// TIA Portal project "pb_slave_test_ZASI_V18" (V18)

(* hardware
DEVICE "S7-1200 station_1"  S7-1200 Station
   slot 0: "Rack_0"  S7-1200 Rack  Rack  V1.0
   slot 1: "PLC_1"  CPU 1212C AC/DC/Rly  6ES7 212-1BE40-0XB0  V4.3
   slot 101: "CM 1243-5"  CM 1243-5  6GK7 243-5DX30-0XE0  V1.3
DEVICE "HMI_1"  KTP700 Basic PN
   slot 0: "HMI_1"  KTP700 Basic PN  6AV2 123-2GB03-0AX0  15.1.0.0
   slot 1: "HMI_RT_1"  KTP700 Basic PN  6AV2 123-2GB03-0AX0  15.1.0.0
   slot 5: "HMI_1.IE_CP_1"  PROFINET Interface  15.0.1.0
      slot 1: "PROFINET Interface_1"  PROFINET Interface
         slot 1: "Port_1"  Port
DEVICE "GSD device_1"  GSD.Device
   slot 0: "Rack_0"  Rail
*)

// ===== PLC "PLC_1"  CPU 1212C AC/DC/Rly =====

VAR_GLOBAL   // PLC tag table "Default tag table"
   "Tag_2" AT %I0.0 : Bool;
   "Tag_1" AT %Q0.0 : Bool;
   "ProfiOut" AT %Q1.0 : "DataRange";
   "System_Byte" AT %MB1 : Byte;
   "FirstScan" AT %M1.0 : Bool;
   "DiagStatusUpdate" AT %M1.1 : Bool;
   "AlwaysTRUE" AT %M1.2 : Bool;
   "AlwaysFALSE" AT %M1.3 : Bool;
   "Clock_Byte" AT %MB0 : Byte;
   "Clock_10Hz" AT %M0.0 : Bool;
   "Clock_5Hz" AT %M0.1 : Bool;
   "Clock_2.5Hz" AT %M0.2 : Bool;
   "Clock_2Hz" AT %M0.3 : Bool;
   "Clock_1.25Hz" AT %M0.4 : Bool;
   "Clock_1Hz" AT %M0.5 : Bool;
   "Clock_0.625Hz" AT %M0.6 : Bool;
   "Clock_0.5Hz" AT %M0.7 : Bool;
   "Length" AT %MD100 : DInt;
   "Length_of_buht" AT %MD104 : DInt;
   "Length_of_buht_current" AT %MD108 : DInt;
   "Velocity" AT %MD112 : DInt;
   "ProfiIn" AT %I1.0 : "DataRange";
   "Dm_pb" AT %ID35 : DWord;
   "Dx_pb" AT %ID39 : UDInt;
   "Dy_pb" AT %ID43 : UDInt;
   "Cx_pb" AT %ID47 : UDInt;
   "Cy_pb" AT %ID51 : UDInt;
   "Error_pb" AT %IB55 : Byte;
   "L_all" AT %ID1 : DInt;
   "set_buht" AT %ID9 : UDInt;
   "L_buht" AT %ID5 : DInt;
   "vel" AT %ID13 : UDInt;
   "Tag_3" AT %QB0 : Byte;
   "Tag_4" AT %QD3 : DInt;
   "ZASI_pb_write_data_addr" AT %QB1 : Byte;
   "Tag_6" AT %QD4 : DInt;
   "Tag_7" AT %QD2 : DInt;
   "ustavka_out" AT %QW6 : Word;
   "proboy" AT %QW4 : Word;
   "reset_length" AT %QB3 : Byte;
   "Ustavka" AT %IW9 : UInt;
   "Voltage" AT %IW13 : UInt;
   "Hi_on" AT %QW2 : UInt;
END_VAR

VAR_GLOBAL   // PLC tag table "global_tags"
   "need_write" AT %M110.0 : Bool;
   "write_addr" AT %MB111 : Byte;
   "new_val" AT %MB112 : Byte;
   "dev_addr" AT %MB113 : Byte;
END_VAR

TYPE "DataRange"
VERSION : 0.1
   STRUCT
      Data : Array[0..36] of Byte;
   END_STRUCT;
END_TYPE

DATA_BLOCK "Zasi_Data"   // DB7
{ S7_Optimized_Access := 'TRUE' }
VERSION : 0.1
   VAR
      Ustavka : Real;
      Capacity : UInt;
      Voltage : Real;
      Hi_on : Byte;
      real_Hi : Byte;
      Proboy : Int;
      write_data_addr : Byte;
      Ustavka_pb : UInt;
      Voltage_pb : UInt;
      Ustavka_HMI : Real;
      Ustavka_HMI_pb : UInt;
      Hi_on_HMI : Byte;
      Ustavka_old_HMI : Real;
      set_Ustavka : Bool;
   END_VAR
BEGIN
END_DATA_BLOCK

// folder: System blocks/Program resources

DATA_BLOCK "IEC_Timer_0_DB"   // DB8
{ S7_Optimized_Access := 'TRUE' }
AUTHOR : Simatic
FAMILY : IEC
NAME : IEC_TMR
VERSION : 1.0
// stored: InstanceOfName IEC_TIMER
"IEC_TIMER"
BEGIN
END_DATA_BLOCK

// folder: (top level)

FUNCTION "Conv_ZASI_data" : Void   // FC3, SCL
{ S7_Optimized_Access := 'TRUE' }
VERSION : 0.1
BEGIN


   "Zasi_Data".Ustavka := UDINT_TO_REAL("Zasi_Data".Ustavka_pb) / 100.0;
   "Zasi_Data".Voltage := UDINT_TO_REAL("Zasi_Data".Voltage_pb) / 100.0;


   "Zasi_Data".Ustavka_HMI_pb := REAL_TO_UDINT("Zasi_Data".Ustavka * 100.0);




   //"Zasi_Data".Ustavka_HMI := "Zasi_Data".Ustavka;


   //"ID_data".pb_HMI_Hi_word := UDINT_TO_WORD(SHR(IN := "ID_data".pb_Set_buht_from_HMI, N := 16));
   //"ID_data".pb_HMI_Low_word := UDINT_TO_WORD("ID_data".pb_Set_buht_from_HMI & 16#FFFF);

   IF "Zasi_Data".Ustavka_old_HMI <> "Zasi_Data".Ustavka_HMI THEN
       "Zasi_Data".set_Ustavka := TRUE;



   END_IF;

   IF ("Zasi_Data".Ustavka_old_HMI = "Zasi_Data".Ustavka_HMI) AND ("Zasi_Data".write_data_addr = 0) THEN
       "Zasi_Data".set_Ustavka := FALSE;
   END_IF;




   IF "Zasi_Data".set_Ustavka  = TRUE THEN

       "Zasi_Data".write_data_addr := 12;
       "Zasi_Data".Ustavka_HMI_pb := REAL_TO_UDINT("Zasi_Data".Ustavka_HMI * 100.0);
   ELSE
       "Zasi_Data".Ustavka_HMI := UDINT_TO_REAL("Zasi_Data".Ustavka_pb) / 100.0;

   END_IF;


   "Zasi_Data".Ustavka_old_HMI := "Zasi_Data".Ustavka_HMI;
END_FUNCTION

ORGANIZATION_BLOCK "Main"   // OB1, LAD, ProgramCycle
TITLE = "Main Program Sweep (Cycle)"
{ S7_Optimized_Access := 'TRUE' }
VERSION : 0.1
   VAR_INPUT
      Initial_Call : Bool;   // Initial call of this OB
      Remanence : Bool;   // =True, if remanent data are available
   END_VAR
BEGIN

REGION Network 1
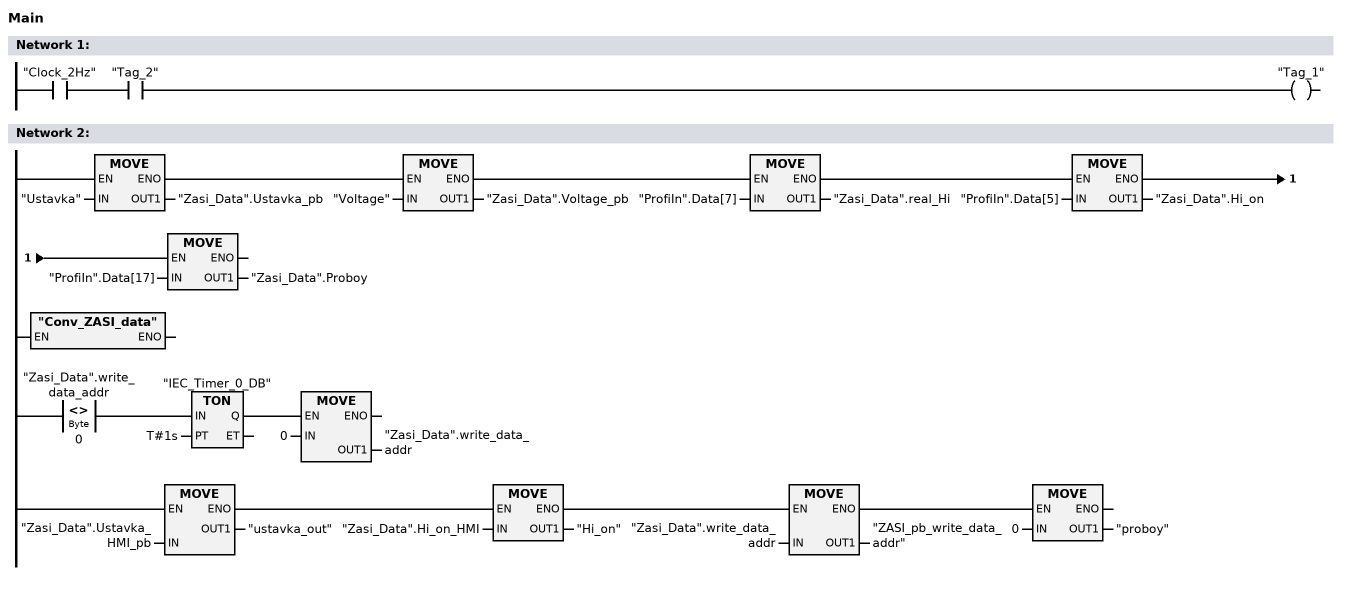
   RUNG wire#powerrail
      Contact( "Clock_2Hz" )
      Contact( "Tag_2" )
      Coil( "Tag_1" )
   END_RUNG
   // the same network as SCL:
   "Tag_1" := "Clock_2Hz" AND "Tag_2";
END_REGION

REGION Network 2
   "Zasi_Data".Ustavka_pb := "Ustavka";
   "Zasi_Data".Voltage_pb := "Voltage";
   "Zasi_Data".real_Hi := "ProfiIn".Data[7];
   "Zasi_Data".Hi_on := "ProfiIn".Data[5];
   "Zasi_Data".Proboy := "ProfiIn".Data[17];
   "Conv_ZASI_data"();
   "IEC_Timer_0_DB".TON(IN := "Zasi_Data".write_data_addr <> 0, PT := T#1s);
   IF "IEC_Timer_0_DB".Q THEN "Zasi_Data".write_data_addr := 0; END_IF;
   "ustavka_out" := "Zasi_Data".Ustavka_HMI_pb;
   "Hi_on" := "Zasi_Data".Hi_on_HMI;
   "ZASI_pb_write_data_addr" := "Zasi_Data".write_data_addr;
   "proboy" := 0;
END_REGION
END_ORGANIZATION_BLOCK

(* ===== HMI "HMI_RT_1" =====
system functions are stored by id; their names below are inferred from use
connection "HMI_Connection_1": ETHERNET, SMART_S7_1200_OMS

HMI tags "Default tag table"
   "need_write" : Bool = PLC need_write AT %M110.0, 1 s
   "write_addr" : Byte = PLC write_addr AT %MB111, 1 s
   "new_val" : Byte = PLC new_val AT %MB112, 1 s
   "dev_addr" : Byte = PLC dev_addr AT %MB113, 1 s
   "Zasi_Data_Voltage" : Real = PLC Zasi_Data.Voltage, 1 s
   "Zasi_Data_Ustavka" : Real = PLC Zasi_Data.Ustavka, 1 s
   "Zasi_Data_Capacity" : UInt = PLC Zasi_Data.Capacity, 1 s
   "Zasi_Data_Proboy" : Int = PLC Zasi_Data.Proboy, 1 s
   "Zasi_Data_Hi_on" : Byte = PLC Zasi_Data.Hi_on, 1 s
   "Zasi_Data_real_Hi" : Byte = PLC Zasi_Data.real_Hi, 1 s
   "Zasi_Data_write_data_addr" : Byte = PLC Zasi_Data.write_data_addr, 1 s
   "Zasi_Data_Ustavka_HMI" : Real = PLC Zasi_Data.Ustavka_HMI, 1 s
   "Zasi_Data_Hi_on_HMI" : Byte = PLC Zasi_Data.Hi_on_HMI, 1 s

text list "LDM_error_messages": 0 ''; 1 'Перекрытие рабочей зоны по двум каналам.'; 2 'Перекрытие верхней границы рабочей зоны по двум каналам'; 3 'Перекрытие нижней границы рабочей зоны по двум каналам'; 4 'Перекрытие нижней границы рабочей зоны по первому каналу'; 5 'Перекрытие верхней границы рабочей зоны по первому каналу'; 6 'Перекрытие рабочей зоны по первому каналу'; 7 'Перекрытие верхней границы рабочей зоны по второму каналу'; 8 'Перекрытие нижней границы рабочей зоны по второму каналу'; 9 'Перекрытие рабочей зоны по второму каналу'; 10 'Перекрытие рабочей зоны по первому каналу и перекрытие верхней границы рабочей зоны по второму каналу'; 11 'Перекрытие рабочей зоны по первому каналу и перекрытие нижней границы рабочей зоны по второму каналу'; 12 'Перекрытие рабочей зоны по второму каналу и перекрытие верхней границы рабочей зоны по первому каналу'; 13 'Перекрытие рабочей зоны по второму каналу и перекрытие нижней границы рабочей зоны по первому каналу'; 14 'Перекрытие верхней границы рабочей зоны по первому каналу и перекрытие нижней границы рабочей зоны по второму каналу'; 15 'Перекрытие нижней границы рабочей зоны по первому каналу и перекрытие верхней границы рабочей зоны по второму каналу'; 16 'Наличие двух и более объектов в зоне измерения'

screen "ZASI" 800x480
   IOField "I/O field_1" at 48,161 size 233x96; FormatPattern 99.99
      ProcessValue <- "Zasi_Data_Voltage"
   IOField "I/O field_2" at 648,163 size 132x96; FormatPattern 99
      ProcessValue <- "Zasi_Data_Proboy"
   IOField "I/O field_3" at 48,379 size 234x96; FormatPattern 99.99
      ProcessValue <- "Zasi_Data_Ustavka_HMI"
   IOField "I/O field_4" at 638,367 size 141x96; FormatPattern 999
      ProcessValue <- "Zasi_Data_Capacity"
   TextField "Text field_1" at 50,101 size 185x62; Text 'Текущее напряжение, кВ'
   TextField "Text field_2" at 641,100 size 133x62; Text 'Количество дефектов'
   TextField "Text field_3" at 45,316 size 185x62; Text 'Испытательное напряжение, кВ'
   TextField "Text field_4" at 635,323 size 139x33; Text 'Емкость, пФ'
   Button "Button_1" at 48,272 size 238x43; TextOff 'Установить'
      on Release: SetTag("Zasi_Data_write_data_addr", 12)
   Button "Button_2" at 646,272 size 135x43; TextOff 'Сброс'
      on Release: SetTag("Zasi_Data_write_data_addr", 16)
   GraphicView "Graphic view_1" at 297,15 size 480x74; Picture "Graphic_1"
   TextField "Text field_5" at 29,0 size 256x100; Text 'Испытатель ЗАСИ'
   Circle "Circle_2" at 424,171 size 82x82
      Appearance <- "Zasi_Data_real_Hi"
   TextField "Text field_6" at 351,115 size 215x33; Text 'Высокое включено'
   Switch "Switch_1" at 376,391 size 204x74; CaptionText 'Switch'; TextOff 'ВЫКЛ'; TextOn 'ВКЛ'
      on Change: SetTag("Zasi_Data_write_data_addr", 10)
      ProcessValue <- "Zasi_Data_Hi_on_HMI"
   TextField "Text field_7" at 365,331 size 212x33; Text 'Включить высокое'
*)